// TIA Portal project "Project maybe not work 1.0" (V17)

(* hardware
DEVICE "S7-1200 station_1"  S7-1200 Station
   slot 0: "Rack_0"  S7-1200 Rack  Rack  V1.0
   slot 1: "PLC_1"  CPU 1214C AC/DC/Rly  6ES7 214-1BG40-0XB0  V4.5
   slot 3: "AQ 1x12BIT_1"  AQ1 signal board  6ES7 232-4HA30-0XB0  V1.0
DEVICE "HMI_1"  TP1500 Comfort
   slot 0: "HMI_1"  TP1500 Comfort  6AV2 124-0QC02-0AX1  17.0.0.0
   slot 1: "HMI_RT_1"  TP1500 Comfort  6AV2 124-0QC02-0AX1  17.0.0.0
   slot 5: "HMI_1.IE_CP_1"  PROFINET Interface  17.0.0.0
      slot 1: "PROFINET Interface_1"  PROFINET Interface
         slot 1: "Port_1"  Port
         slot 2: "Port_2"  Port
   slot 6: "HMI_1.IE_CP_2"  PROFINET Interface  17.0.0.0
      slot 1: "PROFINET Interface_GBit"  PROFINET Interface
         slot 1: "Port_1"  Port
   slot 7: "HMI_1.MPI/DP_CP_1"  MPI/DP Interface  17.0.0.0
*)

// ===== PLC "PLC_1"  CPU 1214C AC/DC/Rly =====

VAR_GLOBAL   // PLC tag table "Default tag table"
   "Tag_1" AT %M40.0 : Bool;
   "Tag_2" AT %M41.0 : Bool;
   "Clock_Byte" AT %MB100 : Byte;
   "Clock_10Hz" AT %M100.0 : Bool;
   "Clock_5Hz" AT %M100.1 : Bool;
   "Clock_2.5Hz" AT %M100.2 : Bool;
   "Clock_2Hz" AT %M100.3 : Bool;
   "Clock_1.25Hz" AT %M100.4 : Bool;
   "Clock_1Hz" AT %M100.5 : Bool;
   "Clock_0.625Hz" AT %M100.6 : Bool;
   "Clock_0.5Hz" AT %M100.7 : Bool;
   "Flash" AT %M36.3 : Bool;
   "Tag_3" AT %MD208 : Real;
   "Tag_4" AT %MD212 : Real;
   "PFC_nodelay" AT %MD218 : Real;
   "Temperature.sp" AT %MW222 : Int;
   "TempDelay" AT %MW226 : Word;
   "Tag_5" AT %MD300 : DWord;
   "Tag_6" AT %MW304 : Word;
END_VAR

VAR_GLOBAL   // PLC tag table "AC_tag_table"
   "QE-200.i" AT %MW64 : Int;   // CO2 ppm(0-1200ppm/ 4-20mA)
   "TFC-201.o" AT %MD80 : Real;   // Intake Air Fan speed(20-100%)
   "PFC-202.o" AT %MD84 : Real;   // Exhaust Air Fan Speed(20-100%)
   "TE-100.i" AT %MW66 : Int;   // Indoor Temperature Sensor (-100 - 100C)
   "TC-101.O" AT %Q0.0 : Bool;   // Heater Control(1=on, 0=off)
   "FCS-110.O" AT %Q0.1 : Bool;   // Intake Damper control(1=open)
   "FCS-111.O" AT %Q0.2 : Bool;   // Intake Damper control (1=closed)
   "FS-113.I" AT %I6.1 : Bool;   // Intake air fan status(1=on)
   "FS-114.I" AT %I7.5 : Bool;   // Intake Damper Closed Status(1=closed)
   "FS-115.I" AT %I7.1 : Bool;   // Intake Damper Open Status(1=open)
   "QE-116.I" AT %I7.3 : Bool;   // Intake vent Smoke Detected(1=smoke in intake vent)
   "FCS-210O" AT %Q0.3 : Bool;   // Exhause Damper control(1=open)
   "FCS-211.O" AT %Q0.4 : Bool;   // Exhaust Damper control(1=closed)
   "FS-212.I" AT %I6.4 : Bool;   // Exhaust air fan status(1=on)
   "FS-213.I" AT %I7.4 : Bool;   // Exhaust Air Damper Closed Status(1=closed)
   "FS-214-I" AT %I7.0 : Bool;   // Exhaust Air Damper Open Status(1=open)
   "FCS-310.O" AT %Q0.5 : Bool;   // Smoke Extraction Fan Control(1=on)
   "FCS-311.O" AT %Q0.6 : Bool;   // Smoke Damper control(1=open)
   "FCS-312.O" AT %Q0.7 : Bool;   // Smoke Damper control(1=closed)
   "FS-313.I" AT %I6.2 : Bool;   // Smoke Fan status(1=on)
   "FS-314.I" AT %I7.2 : Bool;   // Smoke Damper Open Status(1=open)
   "FS-315.I" AT %I7.6 : Bool;   // Smoke Damper Closed Status(1=closed)
   "QE-316.I" AT %I7.7 : Bool;   // Fire Detector(1= no fire, 0=fire)
   "PS-410.I" AT %I6.0 : Bool;   // Start button, rising edge
   "PS-411.I" AT %I6.3 : Bool;   // Stop/Reset button
   "HZ-413.I" AT %I6.5 : Bool;   // Emergency Stop button
   "Setpoint" AT %MD8 : Real;
   "Fire lock" AT %M36.2 : Bool;
   "Start" AT %I4.1 : Bool;
   "Intake Air fan Norm" AT %MD12 : Real;
   "FC" AT %M20.0 : Bool;   // Intake fan control
   "TFC nodelay" AT %MD24 : Real;
   "FC(1)" AT %M20.1 : Bool;   // Exhaust fan control
   "Alarm" AT %M36.0 : Bool;
   "Fire Alarm" AT %M36.1 : Bool;
   "Reset button light" AT %Q1.0 : Bool;
   "Emergency" AT %M36.4 : Bool;
   "QE-200md" AT %MW204 : Word;
   "Co2 Setpoint" AT %MD200 : Real;
   "FanDelay" AT %MW70 : Word;
   "Mitäs Vittus" AT %M2.0 : Bool;
   "Vittus Mitäs" AT %M2.1 : Bool;
END_VAR

DATA_BLOCK "LSim_PT1_DB"   // DB3
{ S7_Optimized_Access := 'TRUE' }
VERSION : 2.01
// stored: InstanceOfName LSim_PT1
"LSim_PT1"
BEGIN
END_DATA_BLOCK

DATA_BLOCK "Many Alarms"   // DB4
{ S7_Optimized_Access := 'FALSE' }
VERSION : 0.1
   VAR
      Alarms : Struct
         "Intake Damper Alarm" : Bool;
         "Fan Alarm" : Bool;
         "Exhaust Damper Alarm" : Bool;
         "Exhaust Fan Alarm" : Bool;
         "Smoke Damper Alarm" : Bool;
         "Smoke Fan Alarm" : Bool;
      END_STRUCT;
   END_VAR
BEGIN
END_DATA_BLOCK

DATA_BLOCK "LSim_Lagging_DB"   // DB5
{ S7_Optimized_Access := 'TRUE' }
VERSION : 2.02
// stored: InstanceOfName LSim_Lagging
"LSim_Lagging"
BEGIN
END_DATA_BLOCK

DATA_BLOCK "Data_Block_Reset_Seq"   // DB6
{ S7_Optimized_Access := 'TRUE' }
VERSION : 0.1
   VAR
      SeqStart : Bool;
      SeqComplete : Bool;
      StepNumber : Int;
      SeqConditions : Array[0..127] of Bool;
      SeqStep : Array[0..127] of Bool;
      SeqTimer_1 : Array[0..127] of TON_TIME;
      SeqTimer : Array[0..127] of TON_TIME;
   END_VAR
BEGIN
END_DATA_BLOCK

DATA_BLOCK "Test"   // DB8
{ S7_Optimized_Access := 'TRUE' }
VERSION : 0.1
   VAR
      "CO2 Level Setpoint" : Int := 0;
      "Temerature Setpoint" : Int;
      "PID TFC Output" : Real;
      "PID TIC Output" : Real;
      "Co2 Input" : Real;
      "TE Input" : Real;
   END_VAR
BEGIN
END_DATA_BLOCK

DATA_BLOCK "Data_Block_Start_Seq"   // DB11
{ S7_Optimized_Access := 'TRUE' }
VERSION : 0.1
   VAR
      SeqStart : Bool;
      SeqComplete : Bool;
      StepNumber : Int;
      SeqConditions : Array[0..127] of Bool;
      SeqStep : Array[0..127] of Bool;
      SeqTimer : Array[0..127] of TON_TIME;
      "To 0" : Bool;
      Start : Bool;
   END_VAR
BEGIN
END_DATA_BLOCK

DATA_BLOCK "Stop_seq_block"   // DB12
{ S7_Optimized_Access := 'TRUE' }
VERSION : 0.1
   VAR
      Sequence_Step : Int;
      SeqStart : Bool;
      SeqComplete : Bool;
      HardwareFailure_CT : Array[0..127] of TON_TIME;
      TimerArray : Array[0..127] of TON_TIME;
   END_VAR
BEGIN
END_DATA_BLOCK

DATA_BLOCK "Fire_Lock_Block"   // DB13
{ S7_Optimized_Access := 'TRUE' }
VERSION : 0.1
   VAR
      Sequence_Step : Int;
      TimerArray : Array[0..127] of TON_TIME;
   END_VAR
BEGIN
END_DATA_BLOCK

DATA_BLOCK "LSim_PT1_DB_1"   // DB16
{ S7_Optimized_Access := 'TRUE' }
VERSION : 2.01
// stored: InstanceOfName LSim_PT1
"LSim_PT1"
BEGIN
END_DATA_BLOCK

DATA_BLOCK "LSim_Lagging_DB_1"   // DB17
{ S7_Optimized_Access := 'TRUE' }
VERSION : 2.02
// stored: InstanceOfName LSim_Lagging
"LSim_Lagging"
BEGIN
END_DATA_BLOCK

DATA_BLOCK "Block_1_DB"   // DB20
{ S7_Optimized_Access := 'TRUE' }
VERSION : 0.1
// stored: InstanceOfName Block_1
"Block_1"
BEGIN
END_DATA_BLOCK

DATA_BLOCK "LSim_PT1_1_DB"   // DB22
{ S7_Optimized_Access := 'TRUE' }
VERSION : 2.01
// stored: InstanceOfName LSim_PT1_1
"LSim_PT1_1"
BEGIN
END_DATA_BLOCK

DATA_BLOCK "LSim_Lagging_1_DB"   // DB23
{ S7_Optimized_Access := 'TRUE' }
VERSION : 2.02
// stored: InstanceOfName LSim_Lagging_1
"LSim_Lagging_1"
BEGIN
END_DATA_BLOCK

DATA_BLOCK "LSim_PT1_DB_2"   // DB25
{ S7_Optimized_Access := 'TRUE' }
VERSION : 2.01
// stored: InstanceOfName LSim_PT1
"LSim_PT1"
BEGIN
END_DATA_BLOCK

DATA_BLOCK "LSim_Lagging_DB_2"   // DB26
{ S7_Optimized_Access := 'TRUE' }
VERSION : 2.02
// stored: InstanceOfName LSim_Lagging
"LSim_Lagging"
BEGIN
END_DATA_BLOCK

DATA_BLOCK "LSim_PT1_DB_3"   // DB28
{ S7_Optimized_Access := 'TRUE' }
VERSION : 2.01
// stored: InstanceOfName LSim_PT1
"LSim_PT1"
BEGIN
END_DATA_BLOCK

DATA_BLOCK "LSim_Lagging_DB_3"   // DB29
{ S7_Optimized_Access := 'TRUE' }
VERSION : 2.02
// stored: InstanceOfName LSim_Lagging
"LSim_Lagging"
BEGIN
END_DATA_BLOCK

// folder: System blocks/Program resources

DATA_BLOCK "IEC_Timer_0_DB"   // DB1
{ S7_Optimized_Access := 'TRUE' }
AUTHOR : Simatic
FAMILY : IEC
NAME : IEC_TMR
VERSION : 1.0
// stored: InstanceOfName IEC_TIMER
"IEC_TIMER"
BEGIN
END_DATA_BLOCK

DATA_BLOCK "IEC_Timer_0_DB_1"   // DB2
{ S7_Optimized_Access := 'TRUE' }
AUTHOR : Simatic
FAMILY : IEC
NAME : IEC_TMR
VERSION : 1.0
// stored: InstanceOfName IEC_TIMER
"IEC_TIMER"
BEGIN
END_DATA_BLOCK

DATA_BLOCK "IEC_Timer_0_DB_4"   // DB9
{ S7_Optimized_Access := 'TRUE' }
AUTHOR : Simatic
FAMILY : IEC
NAME : IEC_TMR
VERSION : 1.0
// stored: InstanceOfName IEC_TIMER
"IEC_TIMER"
BEGIN
END_DATA_BLOCK

DATA_BLOCK "IEC_Timer_0_DB_5"   // DB10
{ S7_Optimized_Access := 'TRUE' }
AUTHOR : Simatic
FAMILY : IEC
NAME : IEC_TMR
VERSION : 1.0
// stored: InstanceOfName IEC_TIMER
"IEC_TIMER"
BEGIN
END_DATA_BLOCK

DATA_BLOCK "IEC_Timer_0_DB_6"   // DB14
{ S7_Optimized_Access := 'TRUE' }
AUTHOR : Simatic
FAMILY : IEC
NAME : IEC_TMR
VERSION : 1.0
// stored: InstanceOfName IEC_TIMER
"IEC_TIMER"
BEGIN
END_DATA_BLOCK

// folder: (top level)

FUNCTION_BLOCK "Block_1"   // FB1, FBD
{ S7_Optimized_Access := 'TRUE' }
VERSION : 0.1
BEGIN

REGION Network 1: Heater Control(1=on, 0=off)
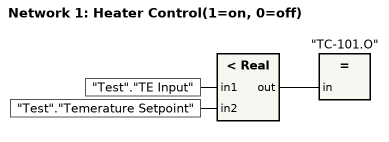
   "TC-101.O" := "Test"."TE Input" < "Test"."Temerature Setpoint";
END_REGION
END_FUNCTION_BLOCK

FUNCTION_BLOCK "LSim_PT1_1"   // FB50, SCL
{ S7_Optimized_Access := 'TRUE' }
VERSION : 2.01
   VAR_INPUT
      calcParam : Bool;   // recalculate with new parameters
      input : Real;   // input signal
      tmLag1 : Real := 1.0;   // time constant T1 [sec]
      gain : Real := 1.0;   // gain factor
      cycle : Real := 0.1;   // cyclic time [sec]
      maxOut : Real := 100.0;   // max. output limit
      minOut : Real;   // min. output limit
      reset : Bool;   // resets all relevant parameters to ‘0’ including the output
   END_VAR
   VAR_OUTPUT
      error : Bool;   // error (#tmLag1 <= 0)
      status : Word;   // status (if #tmLag1 <= 0 then status = 16#8001)
      maxReached : Bool;   // output has reached max. limit
      minReached : Bool;   // output has reached min. limit
      output : Real;   // output signal (if #error = FALSE)
   END_VAR
   VAR
      statRf1 : Real;
      statRe1 : Real;
      statOverfirst : Bool;
      statOutput : Real;
   END_VAR
BEGIN
   //=============================================================================
   //SIEMENS AG
   //(c)Copyright 2017 All Rights Reserved
   //-----------------------------------------------------------------------------
   //Library:       Library for Controlled System Simulation
   //Tested with:   S7-1500 FW V2.0 / S7-1200 FW V4.2
   //Engineering:   STEP 7 V14 Upd2 (TIA Portal)
   //Restrictions:  Cyclic interrupt
   //Requirements:  memory card needed for S7-1500
   //Functionality: Simulation of a PT1-System
   //
   //              gain
   //  F(p) = ---------------
   //          tmLag1 * p + 1
   //          
   //  Call the simulation in a cyclic interrupt with
   //  cyclic interrupt time at least = tmLag1/10!
   //-----------------------------------------------------------------------------
   //Change log table:
   //Version  Date       Expert in charge                Changes applied
   //02.00.00 03.02.2016 Siemens Industry Online Support Release (STEP 7 V13 SP1)
   //02.00.01 02.03.2017 Siemens Industry Online Support Release (STEP 7 V14)
   //=============================================================================
   // check parameter
   IF #tmLag1 <= 0 THEN
     #error := TRUE;
     #status := W#16#8001;     // Parameter Error
     #statOutput := 0;
     #output := 0;
     RETURN;
   ELSE
     #error := FALSE;
     #status := W#16#0000;     // no error
   END_IF;

   IF #calcParam = True OR NOT #statOverfirst THEN
     #statOverfirst:=1;
   // Z-parameters For Laplace PT1-System
   #statRe1 := - EXP(-#cycle/#tmLag1);
   #statRf1 := #gain*(1 + #statRe1);
   END_IF;

   // Differencial Equation of PT1-System
   #statOutput := #input*#statRf1 - #statOutput*#statRe1;

   // max limit of acutating variable
   IF #statOutput > #maxOut THEN
     #statOutput := #maxOut;
     #maxReached:= True;
   ELSE
     #maxReached := False;
   END_IF;

   // min limit of acutating variable
   IF #statOutput < #minOut THEN
     #statOutput := #minOut;
     #minReached := True;
   ELSE
     #minReached := False;
   END_IF;

   IF #reset THEN
     #statOutput := 0;
   END_IF;

   #output := #statOutput;
END_FUNCTION_BLOCK

FUNCTION_BLOCK "LSim_PT1"   // FB51, SCL
{ S7_Optimized_Access := 'TRUE' }
VERSION : 2.01
   VAR_INPUT
      calcParam : Bool;   // recalculate with new parameters
      input : Real;   // input signal
      tmLag1 : Real := 1.0;   // time constant T1 [sec]
      gain : Real := 1.0;   // gain factor
      cycle : Real := 0.1;   // cyclic time [sec]
      maxOut : Real := 100.0;   // max. output limit
      minOut : Real;   // min. output limit
      reset : Bool;   // resets all relevant parameters to ‘0’ including the output
   END_VAR
   VAR_OUTPUT
      error : Bool;   // error (#tmLag1 <= 0)
      status : Word;   // status (if #tmLag1 <= 0 then status = 16#8001)
      maxReached : Bool;   // output has reached max. limit
      minReached : Bool;   // output has reached min. limit
      output : Real;   // output signal (if #error = FALSE)
   END_VAR
   VAR
      statRf1 : Real;
      statRe1 : Real;
      statOverfirst : Bool;
      statOutput : Real;
   END_VAR
BEGIN
   //=============================================================================
   //SIEMENS AG
   //(c)Copyright 2017 All Rights Reserved
   //-----------------------------------------------------------------------------
   //Library:       Library for Controlled System Simulation
   //Tested with:   S7-1500 FW V2.0 / S7-1200 FW V4.2
   //Engineering:   STEP 7 V14 Upd2 (TIA Portal)
   //Restrictions:  Cyclic interrupt
   //Requirements:  memory card needed for S7-1500
   //Functionality: Simulation of a PT1-System
   //
   //              gain
   //  F(p) = ---------------
   //          tmLag1 * p + 1
   //          
   //  Call the simulation in a cyclic interrupt with
   //  cyclic interrupt time at least = tmLag1/10!
   //-----------------------------------------------------------------------------
   //Change log table:
   //Version  Date       Expert in charge                Changes applied
   //02.00.00 03.02.2016 Siemens Industry Online Support Release (STEP 7 V13 SP1)
   //02.00.01 02.03.2017 Siemens Industry Online Support Release (STEP 7 V14)
   //=============================================================================
   // check parameter
   IF #tmLag1 <= 0 THEN
     #error := TRUE;
     #status := W#16#8001;     // Parameter Error
     #statOutput := 0;
     #output := 0;
     RETURN;
   ELSE
     #error := FALSE;
     #status := W#16#0000;     // no error
   END_IF;

   IF #calcParam = True OR NOT #statOverfirst THEN
     #statOverfirst:=1;
   // Z-parameters For Laplace PT1-System
   #statRe1 := - EXP(-#cycle/#tmLag1);
   #statRf1 := #gain*(1 + #statRe1);
   END_IF;

   // Differencial Equation of PT1-System
   #statOutput := #input*#statRf1 - #statOutput*#statRe1;

   // max limit of acutating variable
   IF #statOutput > #maxOut THEN
     #statOutput := #maxOut;
     #maxReached:= True;
   ELSE
     #maxReached := False;
   END_IF;

   // min limit of acutating variable
   IF #statOutput < #minOut THEN
     #statOutput := #minOut;
     #minReached := True;
   ELSE
     #minReached := False;
   END_IF;

   IF #reset THEN
     #statOutput := 0;
   END_IF;

   #output := #statOutput;
END_FUNCTION_BLOCK

FUNCTION_BLOCK "LSim_Lagging"   // FB52, SCL
{ S7_Optimized_Access := 'TRUE' }
VERSION : 2.02
   VAR_INPUT
      input : Real;   // input signal
   END_VAR
   VAR_OUTPUT
      output : Real;   // output signal
   END_VAR
   VAR_IN_OUT
      delayCycles : UInt;   // number of cycles the input signal is delayed (if #delayCycles > #MAX then #delayCycles = #MAX)
   END_VAR
   VAR
      statDelayStore : Array[0..#MAX] of Real;
      statIndexRead : Int;
      statIndexWrite : Int;
   END_VAR
   VAR CONSTANT
      MAX : Int := 100;   // maximum size of array #statDelayStore
   END_VAR
BEGIN
   //=============================================================================
   //SIEMENS AG
   //(c)Copyright 2017 All Rights Reserved
   //-----------------------------------------------------------------------------
   //Library:       Library for Controlled System Simulation
   //Tested with:   S7-1500 FW V2.0 / S7-1200 FW V4.2
   //Engineering:   STEP 7 V14 Upd2 (TIA Portal)
   //Restrictions:  Cyclic interrupt
   //Requirements:  memory card needed for S7-1500
   //Functionality: Simulation of an Tt-System (Lagging)
   //
   //  F(p) = EXP(-p * delayCycles * cyclic interrupt time)
   //          
   //  Call the simulation in a cyclic interrupt with
   //  cyclic interrupt time at least = tmLag1/10!
   //-----------------------------------------------------------------------------
   //Change log table:
   //Version  Date       Expert in charge                Changes applied
   //02.00.00 03.02.2016 Siemens Industry Online Support Release (STEP 7 V13 SP1)
   //02.00.01 02.03.2017 Siemens Industry Online Support Optimize program code
   //02.00.02 02.03.2017 Siemens Industry Online Support Release (STEP 7 V14)
   //=============================================================================

   // Check Parameters
   IF #delayCycles > #MAX THEN
     #delayCycles := INT_TO_UINT(#MAX);
   ELSE
     #delayCycles := #delayCycles;
   END_IF;

   IF #statIndexWrite < #delayCycles THEN
     #statDelayStore[#statIndexWrite] := #input;   // write input at delayStore indexWrite
     #statIndexRead := #statIndexWrite + 1;
     #output := #statDelayStore[#statIndexRead];   // read output from delayStore indexWrite + 1
     #statIndexWrite := #statIndexWrite + 1;       // increment delayStore indexWrite
   ELSE // maximum reached
     #statDelayStore[#statIndexWrite] := #input;   // write input at delayStore maximum
     #statIndexRead := 0;                          // set indexRead to beginning
     #output := #statDelayStore[#statIndexRead];   // read output from delayStore indexRead
     #statIndexWrite := 0;                         // set indexWrite to beginning
   END_IF;
END_FUNCTION_BLOCK

FUNCTION_BLOCK "LSim_Lagging_1"   // FB59, SCL
{ S7_Optimized_Access := 'TRUE' }
VERSION : 2.02
   VAR_INPUT
      input : Real;   // input signal
   END_VAR
   VAR_OUTPUT
      output : Real;   // output signal
   END_VAR
   VAR_IN_OUT
      delayCycles : UInt;   // number of cycles the input signal is delayed (if #delayCycles > #MAX then #delayCycles = #MAX)
   END_VAR
   VAR
      statDelayStore : Array[0..#MAX] of Real;
      statIndexRead : Int;
      statIndexWrite : Int;
   END_VAR
   VAR CONSTANT
      MAX : Int := 100;   // maximum size of array #statDelayStore
   END_VAR
BEGIN
   //=============================================================================
   //SIEMENS AG
   //(c)Copyright 2017 All Rights Reserved
   //-----------------------------------------------------------------------------
   //Library:       Library for Controlled System Simulation
   //Tested with:   S7-1500 FW V2.0 / S7-1200 FW V4.2
   //Engineering:   STEP 7 V14 Upd2 (TIA Portal)
   //Restrictions:  Cyclic interrupt
   //Requirements:  memory card needed for S7-1500
   //Functionality: Simulation of an Tt-System (Lagging)
   //
   //  F(p) = EXP(-p * delayCycles * cyclic interrupt time)
   //          
   //  Call the simulation in a cyclic interrupt with
   //  cyclic interrupt time at least = tmLag1/10!
   //-----------------------------------------------------------------------------
   //Change log table:
   //Version  Date       Expert in charge                Changes applied
   //02.00.00 03.02.2016 Siemens Industry Online Support Release (STEP 7 V13 SP1)
   //02.00.01 02.03.2017 Siemens Industry Online Support Optimize program code
   //02.00.02 02.03.2017 Siemens Industry Online Support Release (STEP 7 V14)
   //=============================================================================

   // Check Parameters
   IF #delayCycles > #MAX THEN
     #delayCycles := INT_TO_UINT(#MAX);
   ELSE
     #delayCycles := #delayCycles;
   END_IF;

   IF #statIndexWrite < #delayCycles THEN
     #statDelayStore[#statIndexWrite] := #input;   // write input at delayStore indexWrite
     #statIndexRead := #statIndexWrite + 1;
     #output := #statDelayStore[#statIndexRead];   // read output from delayStore indexWrite + 1
     #statIndexWrite := #statIndexWrite + 1;       // increment delayStore indexWrite
   ELSE // maximum reached
     #statDelayStore[#statIndexWrite] := #input;   // write input at delayStore maximum
     #statIndexRead := 0;                          // set indexRead to beginning
     #output := #statDelayStore[#statIndexRead];   // read output from delayStore indexRead
     #statIndexWrite := 0;                         // set indexWrite to beginning
   END_IF;
END_FUNCTION_BLOCK

FUNCTION "Reset_Sequence" : Void   // FC1, LAD
{ S7_Optimized_Access := 'TRUE' }
VERSION : 0.1
   VAR_TEMP   // added for the SCL form of the ladder/FBD networks
      _w1 : Bool;
   END_VAR
BEGIN

REGION Network 1: step 1
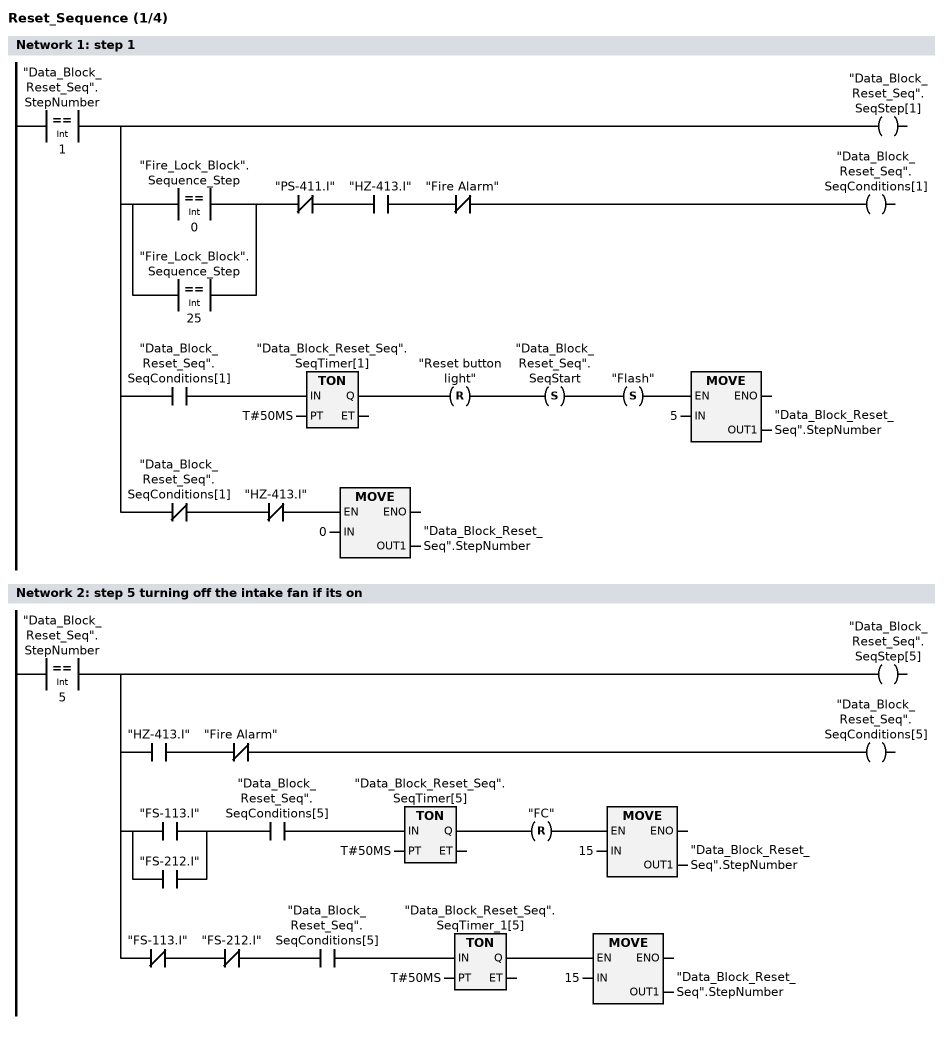
   "Data_Block_Reset_Seq".SeqStep[1] := "Data_Block_Reset_Seq".StepNumber = 1;
   "Data_Block_Reset_Seq".SeqConditions[1] := ("Data_Block_Reset_Seq".StepNumber = 1) AND (("Fire_Lock_Block".Sequence_Step = 0) OR ("Fire_Lock_Block".Sequence_Step = 25)) AND NOT "PS-411.I" AND "HZ-413.I" AND NOT "Fire Alarm";
   "Data_Block_Reset_Seq".SeqTimer[1].TON(IN := ("Data_Block_Reset_Seq".StepNumber = 1) AND "Data_Block_Reset_Seq".SeqConditions[1],
                           PT := T#50MS);
   IF "Data_Block_Reset_Seq".SeqTimer[1].Q THEN
       "Reset button light" := FALSE;
       "Data_Block_Reset_Seq".SeqStart := TRUE;
       "Flash" := TRUE;
   END_IF;
   #_w1 := "Data_Block_Reset_Seq".StepNumber = 1;
   IF "Data_Block_Reset_Seq".SeqTimer[1].Q THEN "Data_Block_Reset_Seq".StepNumber := 5; END_IF;
   IF #_w1 AND NOT "Data_Block_Reset_Seq".SeqConditions[1] AND NOT "HZ-413.I" THEN
       "Data_Block_Reset_Seq".StepNumber := 0;
   END_IF;
END_REGION

REGION Network 2: step 5 turning off the intake fan if its on
   "Data_Block_Reset_Seq".SeqStep[5] := "Data_Block_Reset_Seq".StepNumber = 5;
   "Data_Block_Reset_Seq".SeqConditions[5] := ("Data_Block_Reset_Seq".StepNumber = 5) AND "HZ-413.I" AND NOT "Fire Alarm";
   "Data_Block_Reset_Seq".SeqTimer[5].TON(IN := ("Data_Block_Reset_Seq".StepNumber = 5) AND ("FS-113.I" OR "FS-212.I") AND "Data_Block_Reset_Seq".SeqConditions[5],
                           PT := T#50MS);
   IF "Data_Block_Reset_Seq".SeqTimer[5].Q THEN "FC" := FALSE; END_IF;
   #_w1 := "Data_Block_Reset_Seq".StepNumber = 5;
   IF "Data_Block_Reset_Seq".SeqTimer[5].Q THEN "Data_Block_Reset_Seq".StepNumber := 15; END_IF;
   "Data_Block_Reset_Seq".SeqTimer_1[5].TON(IN := #_w1 AND NOT "FS-113.I" AND NOT "FS-212.I" AND "Data_Block_Reset_Seq".SeqConditions[5],
                           PT := T#50MS);
   IF "Data_Block_Reset_Seq".SeqTimer_1[5].Q THEN "Data_Block_Reset_Seq".StepNumber := 15; END_IF;
END_REGION

REGION Network 3: step 15 Closing the intake damper if its open.
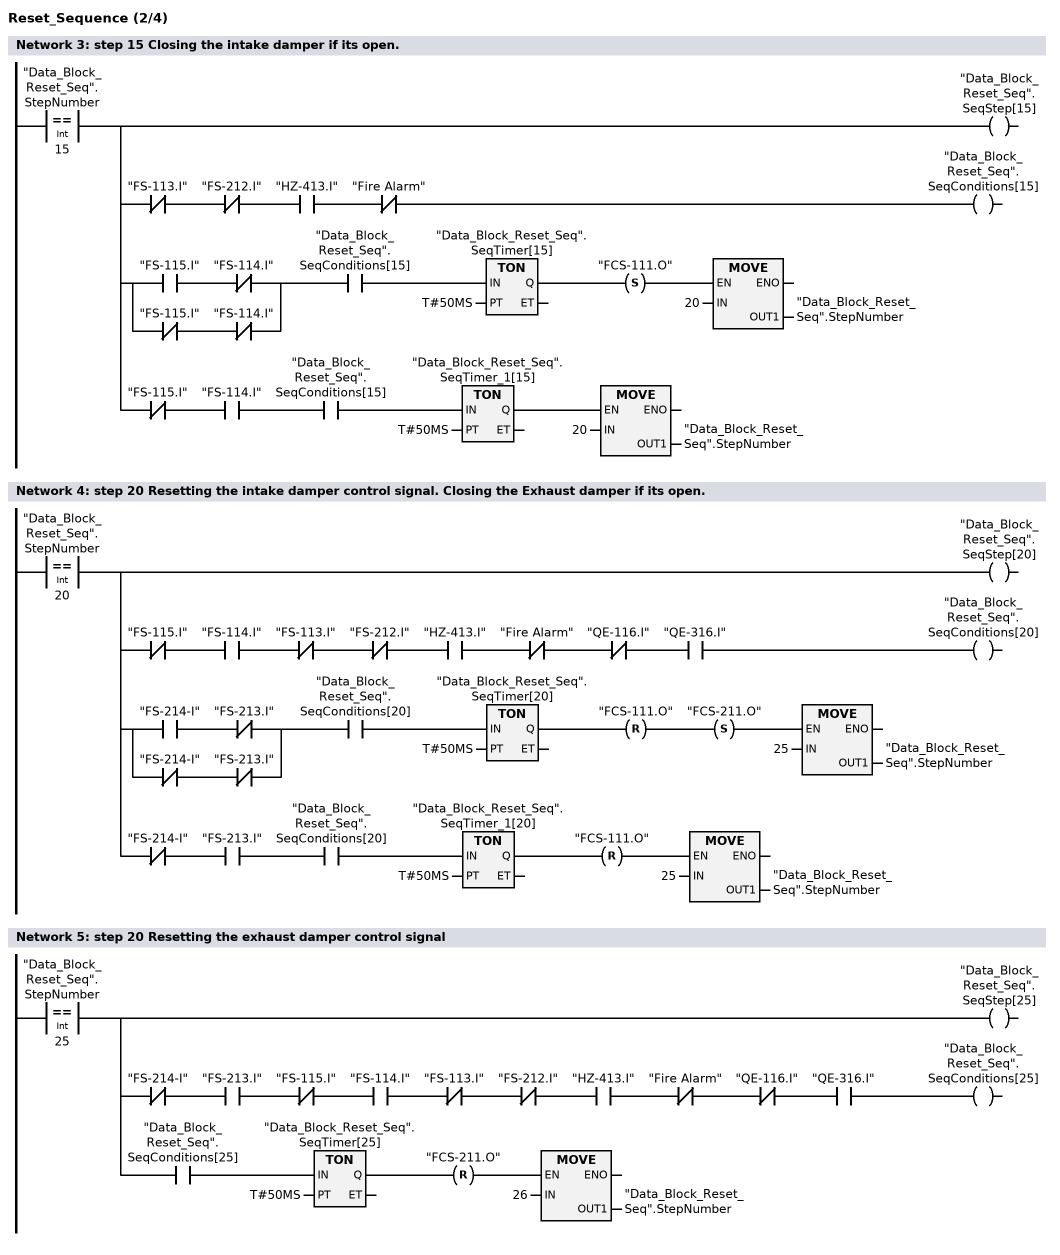
   "Data_Block_Reset_Seq".SeqStep[15] := "Data_Block_Reset_Seq".StepNumber = 15;
   "Data_Block_Reset_Seq".SeqConditions[15] := ("Data_Block_Reset_Seq".StepNumber = 15) AND NOT "FS-113.I" AND NOT "FS-212.I" AND "HZ-413.I" AND NOT "Fire Alarm";
   "Data_Block_Reset_Seq".SeqTimer[15].TON(IN := ("Data_Block_Reset_Seq".StepNumber = 15) AND (("FS-115.I" AND NOT "FS-114.I") OR (NOT "FS-115.I" AND NOT "FS-114.I")) AND "Data_Block_Reset_Seq".SeqConditions[15],
                           PT := T#50MS);
   IF "Data_Block_Reset_Seq".SeqTimer[15].Q THEN "FCS-111.O" := TRUE; END_IF;
   #_w1 := "Data_Block_Reset_Seq".StepNumber = 15;
   IF "Data_Block_Reset_Seq".SeqTimer[15].Q THEN "Data_Block_Reset_Seq".StepNumber := 20; END_IF;
   "Data_Block_Reset_Seq".SeqTimer_1[15].TON(IN := #_w1 AND NOT "FS-115.I" AND "FS-114.I" AND "Data_Block_Reset_Seq".SeqConditions[15],
                           PT := T#50MS);
   IF "Data_Block_Reset_Seq".SeqTimer_1[15].Q THEN "Data_Block_Reset_Seq".StepNumber := 20; END_IF;
END_REGION

REGION Network 4: step 20 Resetting the intake damper control signal. Closing the Exhaust damper if its open.
   "Data_Block_Reset_Seq".SeqStep[20] := "Data_Block_Reset_Seq".StepNumber = 20;
   "Data_Block_Reset_Seq".SeqConditions[20] := ("Data_Block_Reset_Seq".StepNumber = 20) AND NOT "FS-115.I" AND "FS-114.I" AND NOT "FS-113.I" AND NOT "FS-212.I" AND "HZ-413.I" AND NOT "Fire Alarm" AND NOT "QE-116.I" AND "QE-316.I";
   "Data_Block_Reset_Seq".SeqTimer[20].TON(IN := ("Data_Block_Reset_Seq".StepNumber = 20) AND (("FS-214-I" AND NOT "FS-213.I") OR (NOT "FS-214-I" AND NOT "FS-213.I")) AND "Data_Block_Reset_Seq".SeqConditions[20],
                           PT := T#50MS);
   IF "Data_Block_Reset_Seq".SeqTimer[20].Q THEN
       "FCS-111.O" := FALSE;
       "FCS-211.O" := TRUE;
   END_IF;
   #_w1 := "Data_Block_Reset_Seq".StepNumber = 20;
   IF "Data_Block_Reset_Seq".SeqTimer[20].Q THEN "Data_Block_Reset_Seq".StepNumber := 25; END_IF;
   "Data_Block_Reset_Seq".SeqTimer_1[20].TON(IN := #_w1 AND NOT "FS-214-I" AND "FS-213.I" AND "Data_Block_Reset_Seq".SeqConditions[20],
                           PT := T#50MS);
   IF "Data_Block_Reset_Seq".SeqTimer_1[20].Q THEN
       "FCS-111.O" := FALSE;
       "Data_Block_Reset_Seq".StepNumber := 25;
   END_IF;
END_REGION

REGION Network 5: step 20 Resetting the exhaust damper control signal
   "Data_Block_Reset_Seq".SeqStep[25] := "Data_Block_Reset_Seq".StepNumber = 25;
   "Data_Block_Reset_Seq".SeqConditions[25] := ("Data_Block_Reset_Seq".StepNumber = 25) AND NOT "FS-214-I" AND "FS-213.I" AND NOT "FS-115.I" AND "FS-114.I" AND NOT "FS-113.I" AND NOT "FS-212.I" AND "HZ-413.I" AND NOT "Fire Alarm" AND NOT "QE-116.I" AND "QE-316.I";
   "Data_Block_Reset_Seq".SeqTimer[25].TON(IN := ("Data_Block_Reset_Seq".StepNumber = 25) AND "Data_Block_Reset_Seq".SeqConditions[25],
                           PT := T#50MS);
   IF "Data_Block_Reset_Seq".SeqTimer[25].Q THEN
       "FCS-211.O" := FALSE;
       "Data_Block_Reset_Seq".StepNumber := 26;
   END_IF;
END_REGION

REGION Network 6: Step 25 resetting the alarms
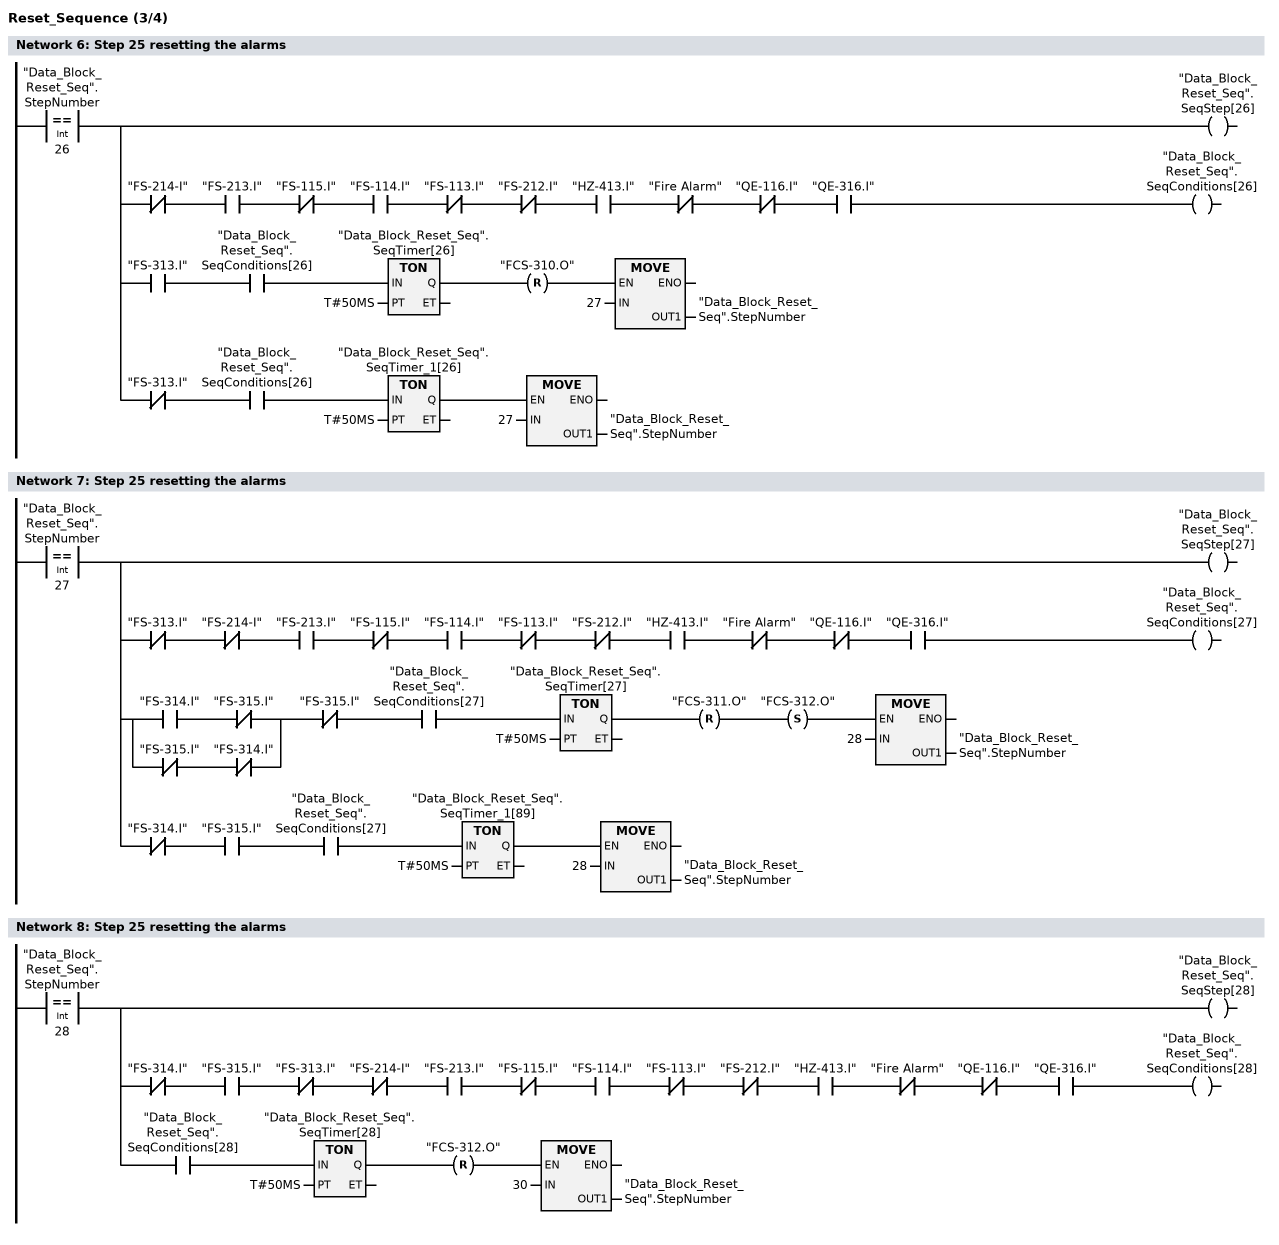
   "Data_Block_Reset_Seq".SeqStep[26] := "Data_Block_Reset_Seq".StepNumber = 26;
   "Data_Block_Reset_Seq".SeqConditions[26] := ("Data_Block_Reset_Seq".StepNumber = 26) AND NOT "FS-214-I" AND "FS-213.I" AND NOT "FS-115.I" AND "FS-114.I" AND NOT "FS-113.I" AND NOT "FS-212.I" AND "HZ-413.I" AND NOT "Fire Alarm" AND NOT "QE-116.I" AND "QE-316.I";
   "Data_Block_Reset_Seq".SeqTimer[26].TON(IN := ("Data_Block_Reset_Seq".StepNumber = 26) AND "FS-313.I" AND "Data_Block_Reset_Seq".SeqConditions[26],
                           PT := T#50MS);
   IF "Data_Block_Reset_Seq".SeqTimer[26].Q THEN "FCS-310.O" := FALSE; END_IF;
   #_w1 := "Data_Block_Reset_Seq".StepNumber = 26;
   IF "Data_Block_Reset_Seq".SeqTimer[26].Q THEN "Data_Block_Reset_Seq".StepNumber := 27; END_IF;
   "Data_Block_Reset_Seq".SeqTimer_1[26].TON(IN := #_w1 AND NOT "FS-313.I" AND "Data_Block_Reset_Seq".SeqConditions[26],
                           PT := T#50MS);
   IF "Data_Block_Reset_Seq".SeqTimer_1[26].Q THEN "Data_Block_Reset_Seq".StepNumber := 27; END_IF;
END_REGION
